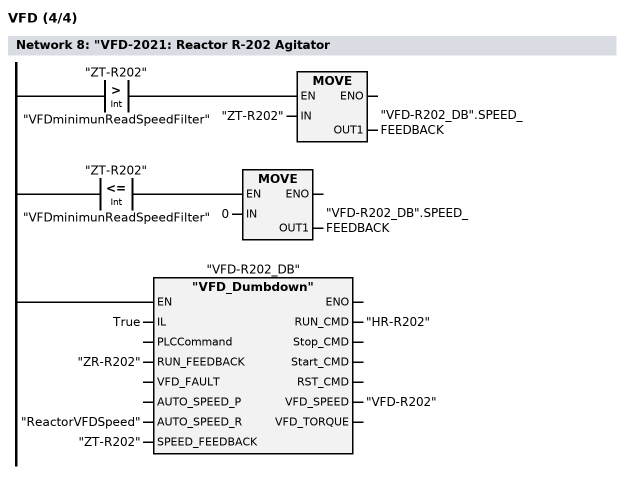
   RUNG wire#powerrail
      { S7_Templates := "SrcType := Int" } GT_Contact(in1 := "ZT-R202", in2 := "VFDminimunReadSpeedFilter")
      { S7_GenerateENO := "TRUE" } Move(in := "ZT-R202", out1 => "VFD-R202_DB".SPEED_FEEDBACK)
   END_RUNG
   RUNG wire#powerrail
      { S7_Templates := "SrcType := Int" } LE_Contact(in1 := "ZT-R202", in2 := "VFDminimunReadSpeedFilter")
      { S7_GenerateENO := "TRUE" } Move(in := 0, out1 => "VFD-R202_DB".SPEED_FEEDBACK)
   END_RUNG
   RUNG wire#powerrail
      "VFD-R202_DB"(IL := True, PLCCommand :=, RUN_FEEDBACK := "ZR-R202", VFD_FAULT :=, AUTO_SPEED_P :=, AUTO_SPEED_R := "ReactorVFDSpeed", SPEED_FEEDBACK := "ZT-R202", RUN_CMD => "HR-R202", Stop_CMD =>, Start_CMD =>, RST_CMD =>, VFD_SPEED => "VFD-R202", VFD_TORQUE =>)
   END_RUNG
   // the same network as SCL:
   IF "ZT-R202" > "VFDminimunReadSpeedFilter" THEN "VFD-R202_DB".SPEED_FEEDBACK := "ZT-R202"; END_IF;
   IF "ZT-R202" <= "VFDminimunReadSpeedFilter" THEN "VFD-R202_DB".SPEED_FEEDBACK := 0; END_IF;
   "VFD-R202_DB"(IL := True,   // "VFD_Dumbdown"
                 RUN_FEEDBACK := "ZR-R202",
                 AUTO_SPEED_R := "ReactorVFDSpeed",
                 SPEED_FEEDBACK := "ZT-R202",
                 RUN_CMD => "HR-R202",
                 VFD_SPEED => "VFD-R202");
END_REGION
END_FUNCTION

// folder: VFD/T103_VFD

FUNCTION "T103_VFD_FC" : Void   // FC112, LAD
{ S7_Optimized_Access := 'TRUE' }
VERSION : 0.1
   VAR_TEMP
      Speed_SP : Real;
   END_VAR
BEGIN

REGION Network 1 (SCL): Speed SP


   IF "VFD-T103_DB".HMI.Controls.Mode = 1 THEN         //Manual Speed SP from HMI

       #Speed_SP := "VFD-T103_DB".HMI.Controls.Speed_Setpoint;

   ELSIF "VFD-T103_DB".HMI.Controls.Mode = 2 THEN      //Auto Speed SP

       #Speed_SP := "T-103_DB".Equipments.VFD."VFD-T103".SP;

   END_IF;

   //Limit the Speed SP
   #Speed_SP := LIMIT_REAL(IN := #Speed_SP, MN := 0.0, MX := 100.0);
END_REGION

REGION Network 2: VFD Profinet Control
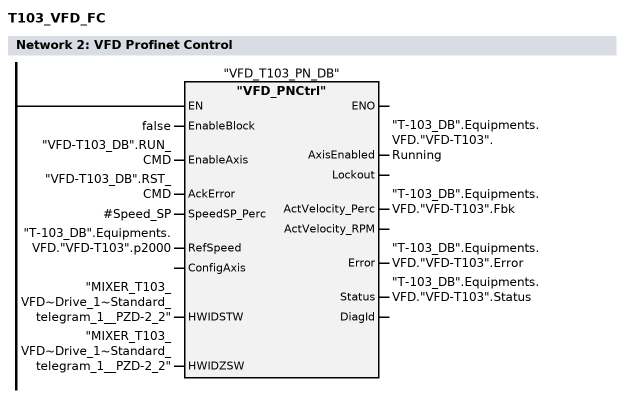
   RUNG wire#powerrail
      "VFD_T103_PN_DB"(EnableBlock := false, EnableAxis := "VFD-T103_DB".RUN_CMD, AckError := "VFD-T103_DB".RST_CMD, SpeedSP_Perc := #Speed_SP, RefSpeed := "T-103_DB".Equipments.VFD."VFD-T103".p2000, ConfigAxis :=, HWIDSTW := "MIXER_T103_VFD~Drive_1~Standard_telegram_1__PZD-2_2", HWIDZSW := "MIXER_T103_VFD~Drive_1~Standard_telegram_1__PZD-2_2", AxisEnabled => "T-103_DB".Equipments.VFD."VFD-T103".Running, Lockout =>, ActVelocity_Perc => "T-103_DB".Equipments.VFD."VFD-T103".Fbk, ActVelocity_RPM =>, Error => "T-103_DB".Equipments.VFD."VFD-T103".Error, Status => "T-103_DB".Equipments.VFD."VFD-T103".Status, DiagId =>)
   END_RUNG
   // the same network as SCL:
   "VFD_T103_PN_DB"(EnableBlock := false,   // "VFD_PNCtrl"
                    EnableAxis := "VFD-T103_DB".RUN_CMD,
                    AckError := "VFD-T103_DB".RST_CMD,
                    SpeedSP_Perc := #Speed_SP,
                    RefSpeed := "T-103_DB".Equipments.VFD."VFD-T103".p2000,
                    HWIDSTW := "MIXER_T103_VFD~Drive_1~Standard_telegram_1__PZD-2_2",
                    HWIDZSW := "MIXER_T103_VFD~Drive_1~Standard_telegram_1__PZD-2_2",
                    AxisEnabled => "T-103_DB".Equipments.VFD."VFD-T103".Running,
                    ActVelocity_Perc => "T-103_DB".Equipments.VFD."VFD-T103".Fbk,
                    Error => "T-103_DB".Equipments.VFD."VFD-T103".Error,
                    Status => "T-103_DB".Equipments.VFD."VFD-T103".Status);
END_REGION
END_FUNCTION

// folder: Valves/Control Valves

FUNCTION "ControlValves" : Void   // FC7, LAD
{ S7_Optimized_Access := 'TRUE' }
VERSION : 0.1
   VAR_TEMP
      BOLL : Bool;
      FEEDBACK : Int;
      OFF : Int;
   END_VAR
BEGIN

REGION Network 1: FV-2011 : T-101 to R-201 Flow Valve
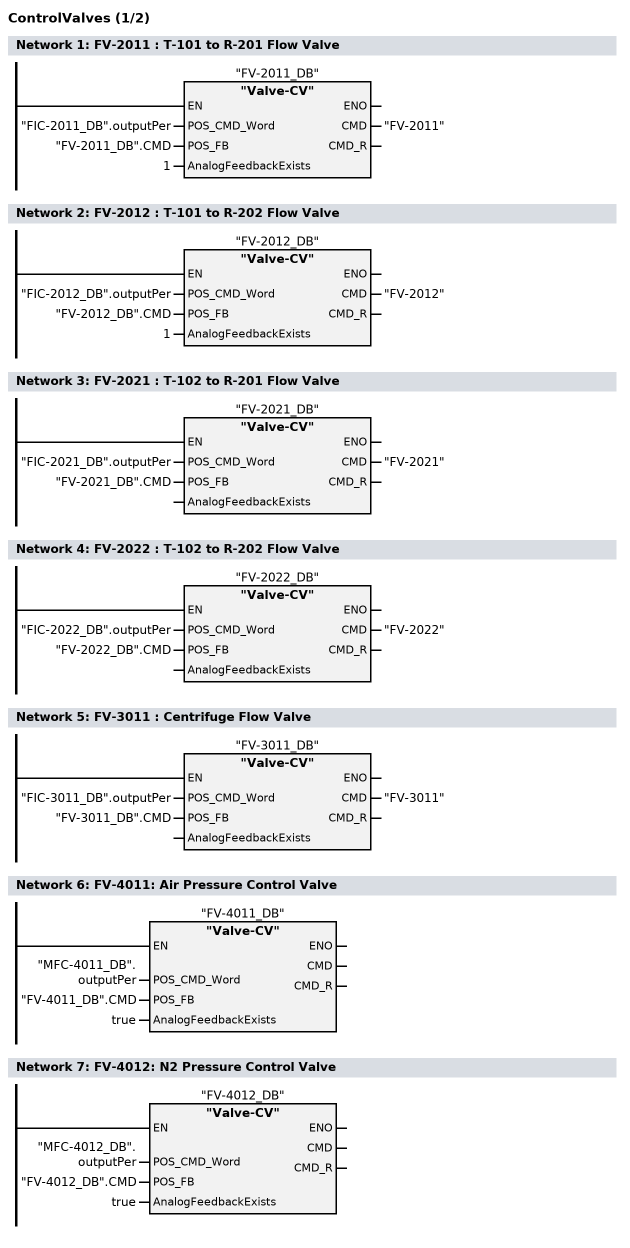
   RUNG wire#powerrail
      "FV-2011_DB"(POS_CMD_Word := "FIC-2011_DB".outputPer, POS_FB := "FV-2011_DB".CMD, AnalogFeedbackExists := 1, CMD => "FV-2011", CMD_R =>)
   END_RUNG
   // the same network as SCL:
   "FV-2011_DB"(POS_CMD_Word := "FIC-2011_DB".outputPer,   // "Valve-CV"
                POS_FB := "FV-2011_DB".CMD,
                AnalogFeedbackExists := 1,
                CMD => "FV-2011");
END_REGION

REGION Network 2: FV-2012 : T-101 to R-202 Flow Valve
   RUNG wire#powerrail
      "FV-2012_DB"(POS_CMD_Word := "FIC-2012_DB".outputPer, POS_FB := "FV-2012_DB".CMD, AnalogFeedbackExists := 1, CMD => "FV-2012", CMD_R =>)
   END_RUNG
   // the same network as SCL:
   "FV-2012_DB"(POS_CMD_Word := "FIC-2012_DB".outputPer,   // "Valve-CV"
                POS_FB := "FV-2012_DB".CMD,
                AnalogFeedbackExists := 1,
                CMD => "FV-2012");
END_REGION

REGION Network 3: FV-2021 : T-102 to R-201 Flow Valve
   RUNG wire#powerrail
      "FV-2021_DB"(POS_CMD_Word := "FIC-2021_DB".outputPer, POS_FB := "FV-2021_DB".CMD, AnalogFeedbackExists :=, CMD => "FV-2021", CMD_R =>)
   END_RUNG
   // the same network as SCL:
   "FV-2021_DB"(POS_CMD_Word := "FIC-2021_DB".outputPer, POS_FB := "FV-2021_DB".CMD, CMD => "FV-2021");   // "Valve-CV"
END_REGION

REGION Network 4: FV-2022 : T-102 to R-202 Flow Valve
   RUNG wire#powerrail
      "FV-2022_DB"(POS_CMD_Word := "FIC-2022_DB".outputPer, POS_FB := "FV-2022_DB".CMD, AnalogFeedbackExists :=, CMD => "FV-2022", CMD_R =>)
   END_RUNG
   // the same network as SCL:
   "FV-2022_DB"(POS_CMD_Word := "FIC-2022_DB".outputPer, POS_FB := "FV-2022_DB".CMD, CMD => "FV-2022");   // "Valve-CV"
END_REGION

REGION Network 5: FV-3011 : Centrifuge Flow Valve
   RUNG wire#powerrail
      "FV-3011_DB"(POS_CMD_Word := "FIC-3011_DB".outputPer, POS_FB := "FV-3011_DB".CMD, AnalogFeedbackExists :=, CMD => "FV-3011", CMD_R =>)
   END_RUNG
   // the same network as SCL:
   "FV-3011_DB"(POS_CMD_Word := "FIC-3011_DB".outputPer, POS_FB := "FV-3011_DB".CMD, CMD => "FV-3011");   // "Valve-CV"
END_REGION

REGION Network 6: FV-4011: Air Pressure Control Valve
   RUNG wire#powerrail
      "FV-4011_DB"(POS_CMD_Word := "MFC-4011_DB".outputPer, POS_FB := "FV-4011_DB".CMD, AnalogFeedbackExists := true, CMD =>, CMD_R =>)
   END_RUNG
   // the same network as SCL:
   "FV-4011_DB"(POS_CMD_Word := "MFC-4011_DB".outputPer,   // "Valve-CV"
                POS_FB := "FV-4011_DB".CMD,
                AnalogFeedbackExists := true);
END_REGION

REGION Network 7: FV-4012: N2 Pressure Control Valve
   RUNG wire#powerrail
      "FV-4012_DB"(POS_CMD_Word := "MFC-4012_DB".outputPer, POS_FB := "FV-4012_DB".CMD, AnalogFeedbackExists := true, CMD =>, CMD_R =>)
   END_RUNG
   // the same network as SCL:
   "FV-4012_DB"(POS_CMD_Word := "MFC-4012_DB".outputPer,   // "Valve-CV"
                POS_FB := "FV-4012_DB".CMD,
                AnalogFeedbackExists := true);
END_REGION

REGION Network 8: FV-4021: Pressure Control Valve
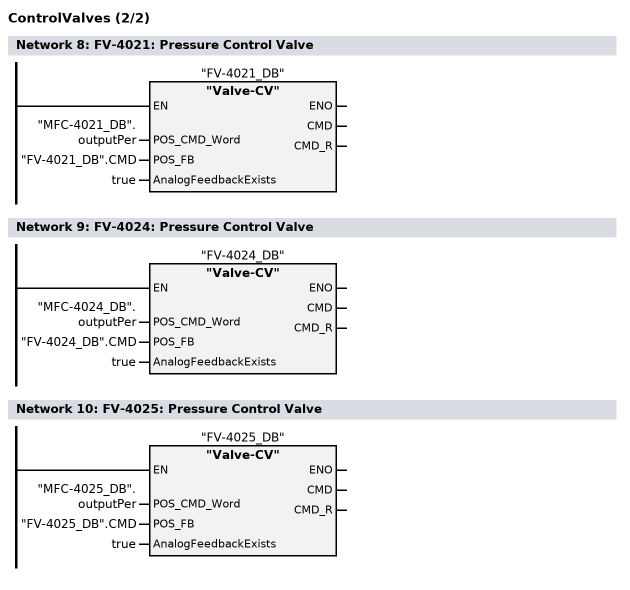
   RUNG wire#powerrail
      "FV-4021_DB"(POS_CMD_Word := "MFC-4021_DB".outputPer, POS_FB := "FV-4021_DB".CMD, AnalogFeedbackExists := true, CMD =>, CMD_R =>)
   END_RUNG
   // the same network as SCL:
   "FV-4021_DB"(POS_CMD_Word := "MFC-4021_DB".outputPer,   // "Valve-CV"
                POS_FB := "FV-4021_DB".CMD,
                AnalogFeedbackExists := true);
END_REGION

REGION Network 9: FV-4024: Pressure Control Valve
   RUNG wire#powerrail
      "FV-4024_DB"(POS_CMD_Word := "MFC-4024_DB".outputPer, POS_FB := "FV-4024_DB".CMD, AnalogFeedbackExists := true, CMD =>, CMD_R =>)
   END_RUNG
   // the same network as SCL:
   "FV-4024_DB"(POS_CMD_Word := "MFC-4024_DB".outputPer,   // "Valve-CV"
                POS_FB := "FV-4024_DB".CMD,
                AnalogFeedbackExists := true);
END_REGION

REGION Network 10: FV-4025: Pressure Control Valve
   RUNG wire#powerrail
      "FV-4025_DB"(POS_CMD_Word := "MFC-4025_DB".outputPer, POS_FB := "FV-4025_DB".CMD, AnalogFeedbackExists := true, CMD =>, CMD_R =>)
   END_RUNG
   // the same network as SCL:
   "FV-4025_DB"(POS_CMD_Word := "MFC-4025_DB".outputPer,   // "Valve-CV"
                POS_FB := "FV-4025_DB".CMD,
                AnalogFeedbackExists := true);
END_REGION
END_FUNCTION

// folder: Valves/Solenoid Valve

FUNCTION "SolenoidValve" : Void   // FC2, LAD
{ S7_Optimized_Access := 'TRUE' }
VERSION : 0.1
BEGIN

REGION Network 1: XV-1041 : T-101 Water Valve
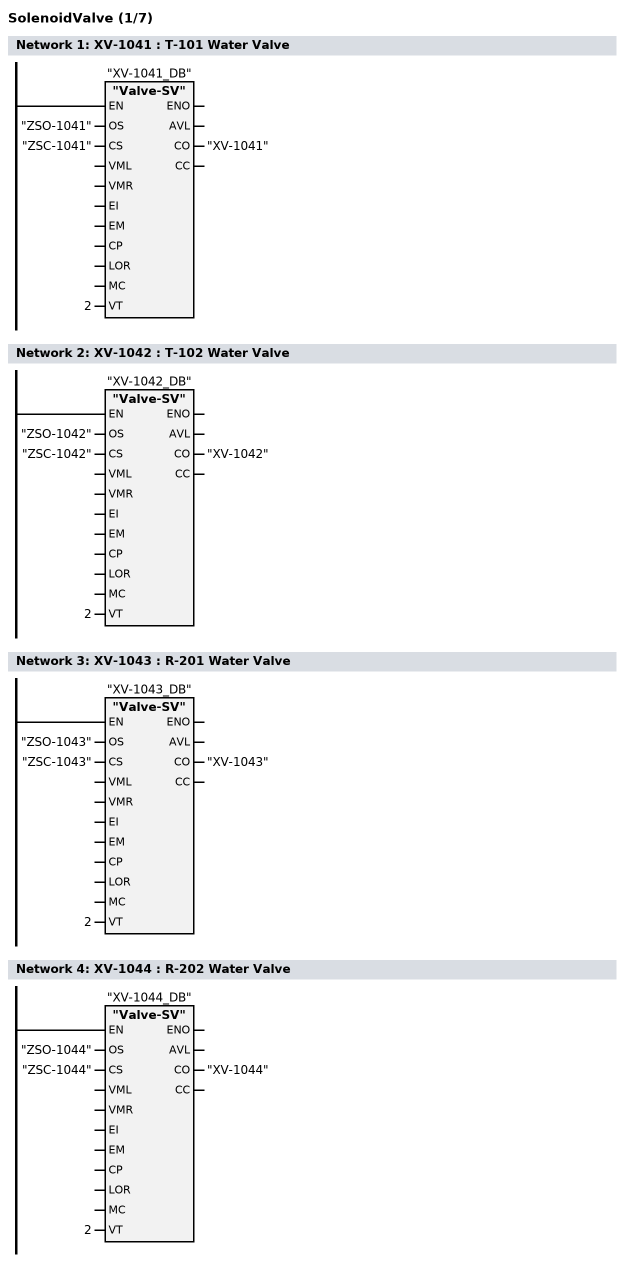
   RUNG wire#powerrail
      "XV-1041_DB"(OS := "ZSO-1041", CS := "ZSC-1041", VML :=, VMR :=, EI :=, EM :=, CP :=, LOR :=, MC :=, VT := 2, AVL =>, CO => "XV-1041", CC =>)
   END_RUNG
   // the same network as SCL:
   "XV-1041_DB"(OS := "ZSO-1041", CS := "ZSC-1041", VT := 2, CO => "XV-1041");   // "Valve-SV"
END_REGION

REGION Network 2: XV-1042 : T-102 Water Valve
   RUNG wire#powerrail
      "XV-1042_DB"(OS := "ZSO-1042", CS := "ZSC-1042", VML :=, VMR :=, EI :=, EM :=, CP :=, LOR :=, MC :=, VT := 2, AVL =>, CO => "XV-1042", CC =>)
   END_RUNG
   // the same network as SCL:
   "XV-1042_DB"(OS := "ZSO-1042", CS := "ZSC-1042", VT := 2, CO => "XV-1042");   // "Valve-SV"
END_REGION

REGION Network 3: XV-1043 : R-201 Water Valve
   RUNG wire#powerrail
      "XV-1043_DB"(OS := "ZSO-1043", CS := "ZSC-1043", VML :=, VMR :=, EI :=, EM :=, CP :=, LOR :=, MC :=, VT := 2, AVL =>, CO => "XV-1043", CC =>)
   END_RUNG
   // the same network as SCL:
   "XV-1043_DB"(OS := "ZSO-1043", CS := "ZSC-1043", VT := 2, CO => "XV-1043");   // "Valve-SV"
END_REGION

REGION Network 4: XV-1044 : R-202 Water Valve
   RUNG wire#powerrail
      "XV-1044_DB"(OS := "ZSO-1044", CS := "ZSC-1044", VML :=, VMR :=, EI :=, EM :=, CP :=, LOR :=, MC :=, VT := 2, AVL =>, CO => "XV-1044", CC =>)
   END_RUNG
   // the same network as SCL:
   "XV-1044_DB"(OS := "ZSO-1044", CS := "ZSC-1044", VT := 2, CO => "XV-1044");   // "Valve-SV"
END_REGION

REGION Network 5: XV-1045 : C-301 Water Valve
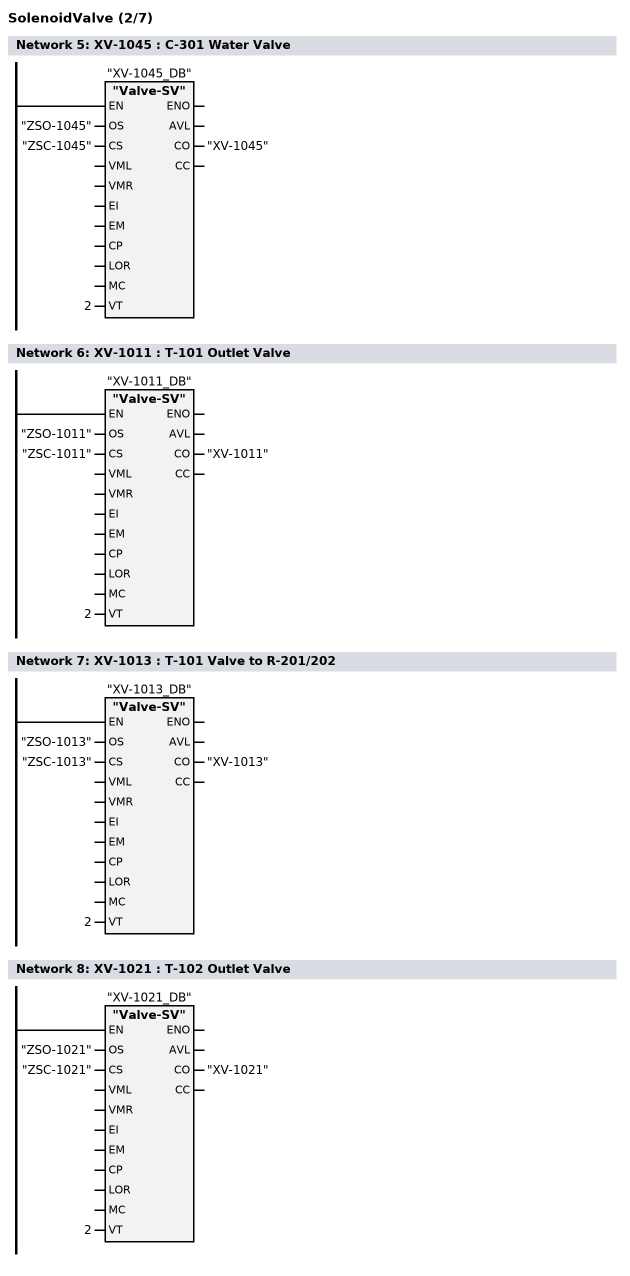
   RUNG wire#powerrail
      "XV-1045_DB"(OS := "ZSO-1045", CS := "ZSC-1045", VML :=, VMR :=, EI :=, EM :=, CP :=, LOR :=, MC :=, VT := 2, AVL =>, CO => "XV-1045", CC =>)
   END_RUNG
   // the same network as SCL:
   "XV-1045_DB"(OS := "ZSO-1045", CS := "ZSC-1045", VT := 2, CO => "XV-1045");   // "Valve-SV"
END_REGION

REGION Network 6: XV-1011 : T-101 Outlet Valve
   RUNG wire#powerrail
      "XV-1011_DB"(OS := "ZSO-1011", CS := "ZSC-1011", VML :=, VMR :=, EI :=, EM :=, CP :=, LOR :=, MC :=, VT := 2, AVL =>, CO => "XV-1011", CC =>)
   END_RUNG
   // the same network as SCL:
   "XV-1011_DB"(OS := "ZSO-1011", CS := "ZSC-1011", VT := 2, CO => "XV-1011");   // "Valve-SV"
END_REGION

REGION Network 7: XV-1013 : T-101 Valve to R-201/202
   RUNG wire#powerrail
      "XV-1013_DB"(OS := "ZSO-1013", CS := "ZSC-1013", VML :=, VMR :=, EI :=, EM :=, CP :=, LOR :=, MC :=, VT := 2, AVL =>, CO => "XV-1013", CC =>)
   END_RUNG
   // the same network as SCL:
   "XV-1013_DB"(OS := "ZSO-1013", CS := "ZSC-1013", VT := 2, CO => "XV-1013");   // "Valve-SV"
END_REGION

REGION Network 8: XV-1021 : T-102 Outlet Valve
   RUNG wire#powerrail
      "XV-1021_DB"(OS := "ZSO-1021", CS := "ZSC-1021", VML :=, VMR :=, EI :=, EM :=, CP :=, LOR :=, MC :=, VT := 2, AVL =>, CO => "XV-1021", CC =>)
   END_RUNG
   // the same network as SCL:
   "XV-1021_DB"(OS := "ZSO-1021", CS := "ZSC-1021", VT := 2, CO => "XV-1021");   // "Valve-SV"
END_REGION

REGION Network 9: XV-1023 : T-102 valve to R-201/202
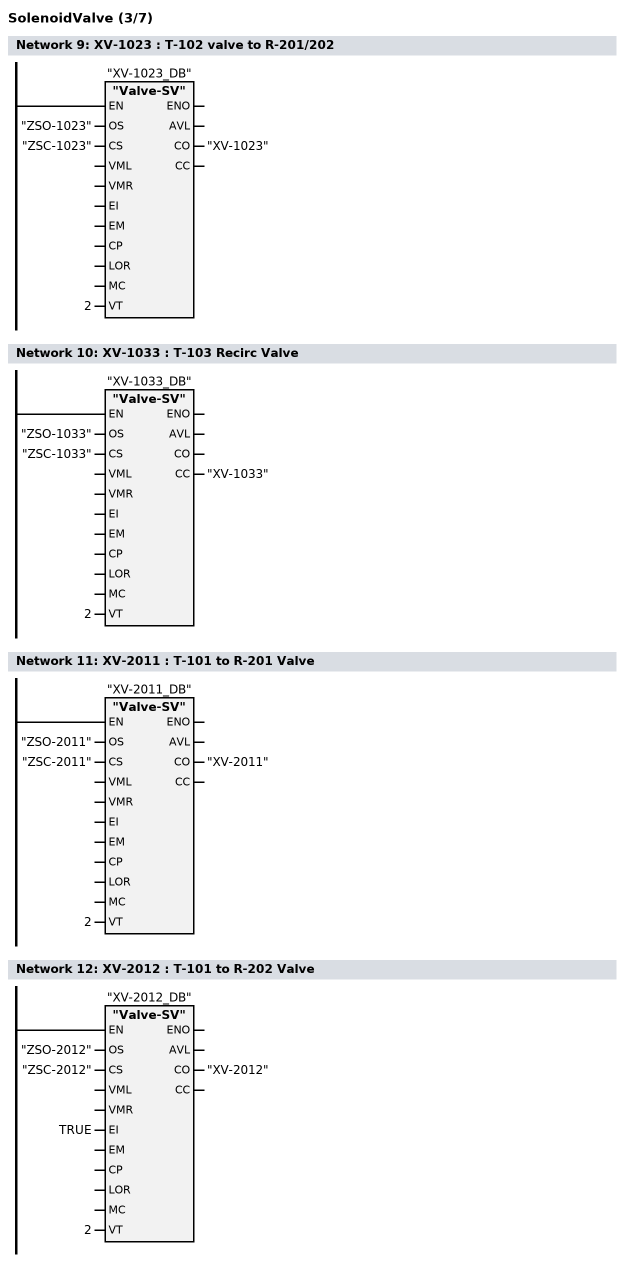
   RUNG wire#powerrail
      "XV-1023_DB"(OS := "ZSO-1023", CS := "ZSC-1023", VML :=, VMR :=, EI :=, EM :=, CP :=, LOR :=, MC :=, VT := 2, AVL =>, CO => "XV-1023", CC =>)
   END_RUNG
   // the same network as SCL:
   "XV-1023_DB"(OS := "ZSO-1023", CS := "ZSC-1023", VT := 2, CO => "XV-1023");   // "Valve-SV"
END_REGION

REGION Network 10: XV-1033 : T-103 Recirc Valve
   RUNG wire#powerrail
      "XV-1033_DB"(OS := "ZSO-1033", CS := "ZSC-1033", VML :=, VMR :=, EI :=, EM :=, CP :=, LOR :=, MC :=, VT := 2, AVL =>, CO =>, CC => "XV-1033")
   END_RUNG
   // the same network as SCL:
   "XV-1033_DB"(OS := "ZSO-1033", CS := "ZSC-1033", VT := 2, CC => "XV-1033");   // "Valve-SV"
END_REGION

REGION Network 11: XV-2011 : T-101 to R-201 Valve
   RUNG wire#powerrail
      "XV-2011_DB"(OS := "ZSO-2011", CS := "ZSC-2011", VML :=, VMR :=, EI :=, EM :=, CP :=, LOR :=, MC :=, VT := 2, AVL =>, CO => "XV-2011", CC =>)
   END_RUNG
   // the same network as SCL:
   "XV-2011_DB"(OS := "ZSO-2011", CS := "ZSC-2011", VT := 2, CO => "XV-2011");   // "Valve-SV"
END_REGION

REGION Network 12: XV-2012 : T-101 to R-202 Valve
   RUNG wire#powerrail
      "XV-2012_DB"(OS := "ZSO-2012", CS := "ZSC-2012", VML :=, VMR :=, EI := TRUE, EM :=, CP :=, LOR :=, MC :=, VT := 2, AVL =>, CO => "XV-2012", CC =>)
   END_RUNG
   // the same network as SCL:
   "XV-2012_DB"(OS := "ZSO-2012", CS := "ZSC-2012", EI := TRUE, VT := 2, CO => "XV-2012");   // "Valve-SV"
END_REGION

REGION Network 13: XV-2021 : T-102 to R-201 Valve
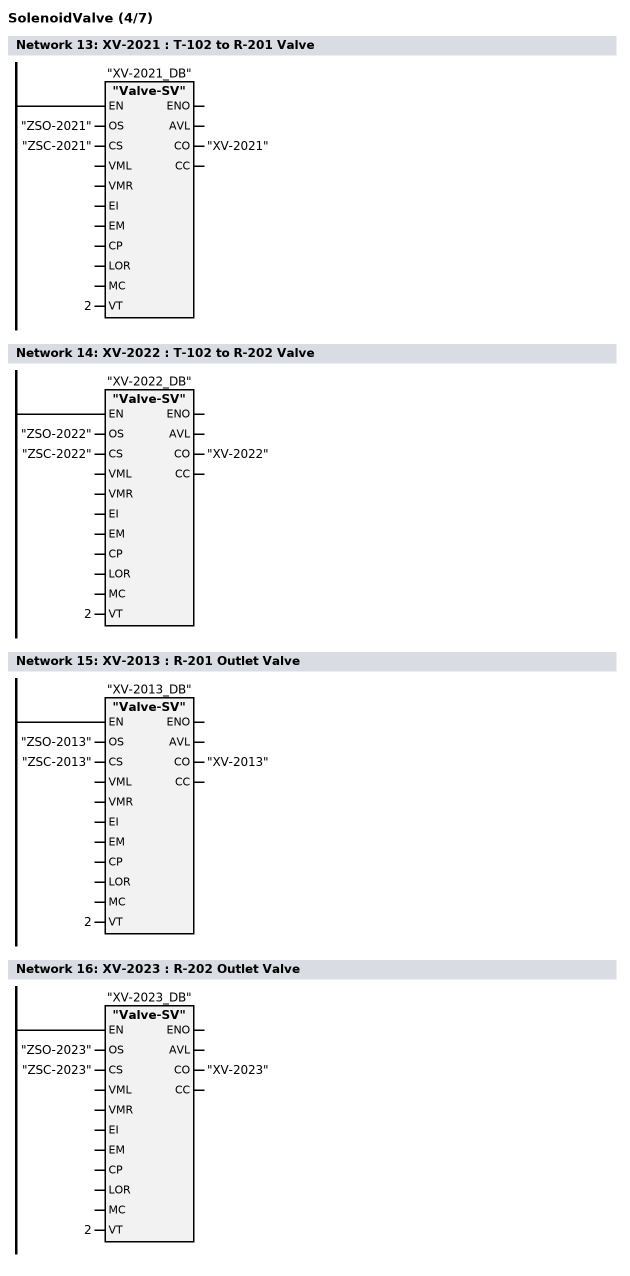
   RUNG wire#powerrail
      "XV-2021_DB"(OS := "ZSO-2021", CS := "ZSC-2021", VML :=, VMR :=, EI :=, EM :=, CP :=, LOR :=, MC :=, VT := 2, AVL =>, CO => "XV-2021", CC =>)
   END_RUNG
   // the same network as SCL:
   "XV-2021_DB"(OS := "ZSO-2021", CS := "ZSC-2021", VT := 2, CO => "XV-2021");   // "Valve-SV"
END_REGION

REGION Network 14: XV-2022 : T-102 to R-202 Valve
   RUNG wire#powerrail
      "XV-2022_DB"(OS := "ZSO-2022", CS := "ZSC-2022", VML :=, VMR :=, EI :=, EM :=, CP :=, LOR :=, MC :=, VT := 2, AVL =>, CO => "XV-2022", CC =>)
   END_RUNG
   // the same network as SCL:
   "XV-2022_DB"(OS := "ZSO-2022", CS := "ZSC-2022", VT := 2, CO => "XV-2022");   // "Valve-SV"
END_REGION

REGION Network 15: XV-2013 : R-201 Outlet Valve
   RUNG wire#powerrail
      "XV-2013_DB"(OS := "ZSO-2013", CS := "ZSC-2013", VML :=, VMR :=, EI :=, EM :=, CP :=, LOR :=, MC :=, VT := 2, AVL =>, CO => "XV-2013", CC =>)
   END_RUNG
   // the same network as SCL:
   "XV-2013_DB"(OS := "ZSO-2013", CS := "ZSC-2013", VT := 2, CO => "XV-2013");   // "Valve-SV"
END_REGION

REGION Network 16: XV-2023 : R-202 Outlet Valve
   RUNG wire#powerrail
      "XV-2023_DB"(OS := "ZSO-2023", CS := "ZSC-2023", VML :=, VMR :=, EI :=, EM :=, CP :=, LOR :=, MC :=, VT := 2, AVL =>, CO => "XV-2023", CC =>)
   END_RUNG
   // the same network as SCL:
   "XV-2023_DB"(OS := "ZSO-2023", CS := "ZSC-2023", VT := 2, CO => "XV-2023");   // "Valve-SV"
END_REGION

REGION Network 17: XV-1031 : R-201/202 to T-103 Valve
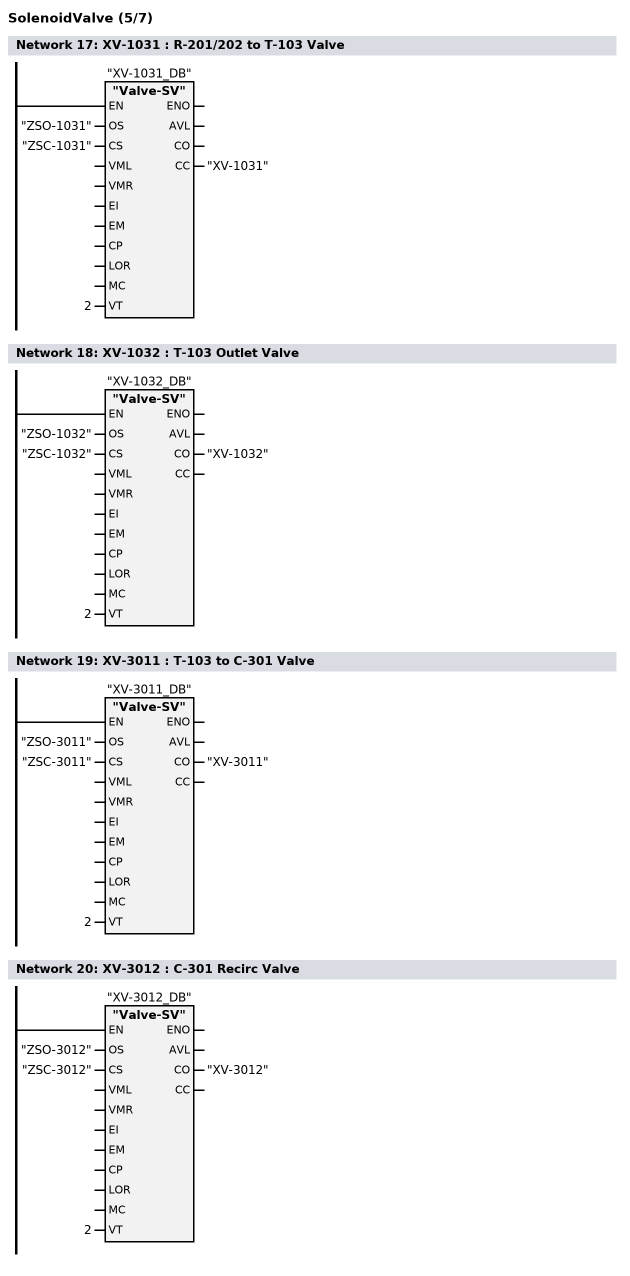
   RUNG wire#powerrail
      "XV-1031_DB"(OS := "ZSO-1031", CS := "ZSC-1031", VML :=, VMR :=, EI :=, EM :=, CP :=, LOR :=, MC :=, VT := 2, AVL =>, CO =>, CC => "XV-1031")
   END_RUNG
   // the same network as SCL:
   "XV-1031_DB"(OS := "ZSO-1031", CS := "ZSC-1031", VT := 2, CC => "XV-1031");   // "Valve-SV"
END_REGION

REGION Network 18: XV-1032 : T-103 Outlet Valve
   RUNG wire#powerrail
      "XV-1032_DB"(OS := "ZSO-1032", CS := "ZSC-1032", VML :=, VMR :=, EI :=, EM :=, CP :=, LOR :=, MC :=, VT := 2, AVL =>, CO => "XV-1032", CC =>)
   END_RUNG
   // the same network as SCL:
   "XV-1032_DB"(OS := "ZSO-1032", CS := "ZSC-1032", VT := 2, CO => "XV-1032");   // "Valve-SV"
END_REGION

REGION Network 19: XV-3011 : T-103 to C-301 Valve
   RUNG wire#powerrail
      "XV-3011_DB"(OS := "ZSO-3011", CS := "ZSC-3011", VML :=, VMR :=, EI :=, EM :=, CP :=, LOR :=, MC :=, VT := 2, AVL =>, CO => "XV-3011", CC =>)
   END_RUNG
   // the same network as SCL:
   "XV-3011_DB"(OS := "ZSO-3011", CS := "ZSC-3011", VT := 2, CO => "XV-3011");   // "Valve-SV"
END_REGION

REGION Network 20: XV-3012 : C-301 Recirc Valve
   RUNG wire#powerrail
      "XV-3012_DB"(OS := "ZSO-3012", CS := "ZSC-3012", VML :=, VMR :=, EI :=, EM :=, CP :=, LOR :=, MC :=, VT := 2, AVL =>, CO => "XV-3012", CC =>)
   END_RUNG
   // the same network as SCL:
   "XV-3012_DB"(OS := "ZSO-3012", CS := "ZSC-3012", VT := 2, CO => "XV-3012");   // "Valve-SV"
END_REGION

REGION Network 21: XV-3013 : C-301 to ST-301 Valve
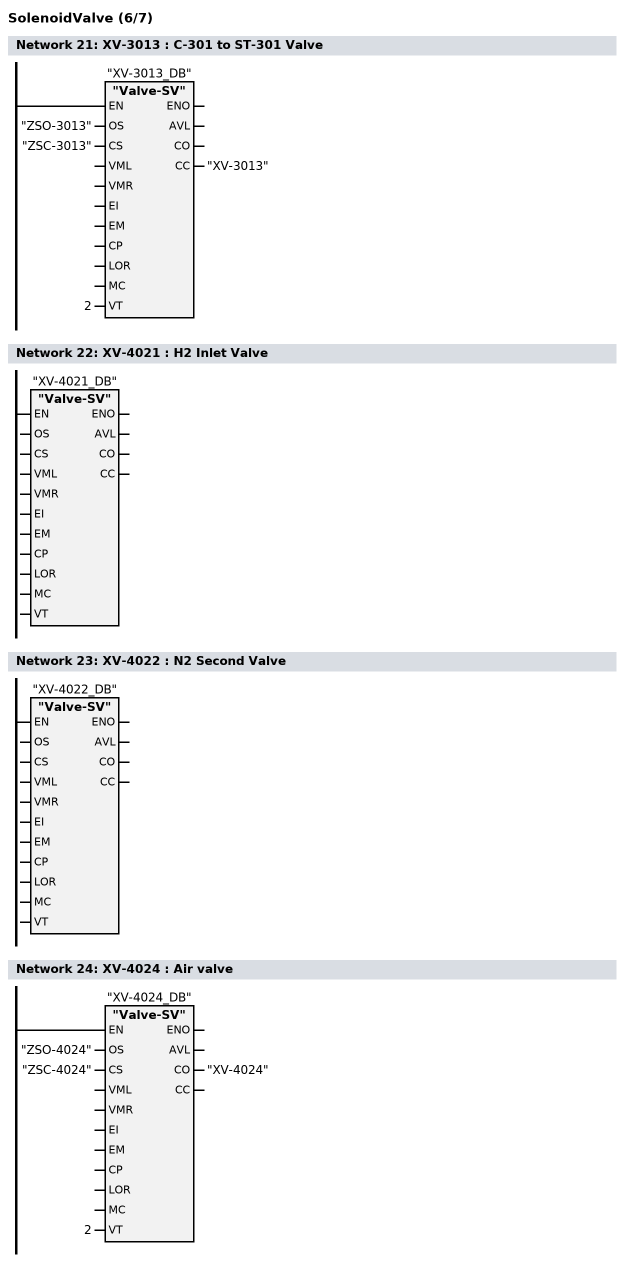
   RUNG wire#powerrail
      "XV-3013_DB"(OS := "ZSO-3013", CS := "ZSC-3013", VML :=, VMR :=, EI :=, EM :=, CP :=, LOR :=, MC :=, VT := 2, AVL =>, CO =>, CC => "XV-3013")
   END_RUNG
   // the same network as SCL:
   "XV-3013_DB"(OS := "ZSO-3013", CS := "ZSC-3013", VT := 2, CC => "XV-3013");   // "Valve-SV"
END_REGION

REGION Network 22: XV-4021 : H2 Inlet Valve
   RUNG wire#powerrail
      "XV-4021_DB"(OS :=, CS :=, VML :=, VMR :=, EI :=, EM :=, CP :=, LOR :=, MC :=, VT :=, AVL =>, CO =>, CC =>)
   END_RUNG
   // the same network as SCL:
   "XV-4021_DB"();   // "Valve-SV"
END_REGION

REGION Network 23: XV-4022 : N2 Second Valve
   RUNG wire#powerrail
      "XV-4022_DB"(OS :=, CS :=, VML :=, VMR :=, EI :=, EM :=, CP :=, LOR :=, MC :=, VT :=, AVL =>, CO =>, CC =>)
   END_RUNG
   // the same network as SCL:
   "XV-4022_DB"();   // "Valve-SV"
END_REGION

REGION Network 24: XV-4024 : Air valve
   RUNG wire#powerrail
      "XV-4024_DB"(OS := "ZSO-4024", CS := "ZSC-4024", VML :=, VMR :=, EI :=, EM :=, CP :=, LOR :=, MC :=, VT := 2, AVL =>, CO => "XV-4024", CC =>)
   END_RUNG
   // the same network as SCL:
   "XV-4024_DB"(OS := "ZSO-4024", CS := "ZSC-4024", VT := 2, CO => "XV-4024");   // "Valve-SV"
END_REGION

REGION Network 25: XV-4025 : N2 Air valve
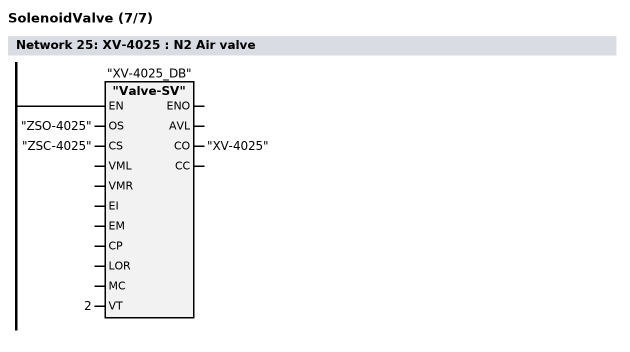
   RUNG wire#powerrail
      "XV-4025_DB"(OS := "ZSO-4025", CS := "ZSC-4025", VML :=, VMR :=, EI :=, EM :=, CP :=, LOR :=, MC :=, VT := 2, AVL =>, CO => "XV-4025", CC =>)
   END_RUNG
   // the same network as SCL:
   "XV-4025_DB"(OS := "ZSO-4025", CS := "ZSC-4025", VT := 2, CO => "XV-4025");   // "Valve-SV"
END_REGION
END_FUNCTION